VERSION : 0.0
   STRUCT
      Config_bit_Converter : Bool;   // Configuration with frequency converter
      Config_bit_Converter_SW : Bool;   // Configuration with frequency converter with Set value
      Config_bit_Heating_ON : Bool;
      config_bit_Heating_Int : Bool;
      Config_bit_Cooling_ON : Bool;
      Config_bit_Cooling_Int : Bool;
      Config_bit_Filling_ON : Bool;
      Config_bit_Filling_Int : Bool;
      Config_bit_Charging_ON : Bool;
      Config_bit_Charging_Int : Bool;
      RunTime : S5Time;
      PauseTime : S5Time;
   END_STRUCT;
END_TYPE

TYPE "UDT102_RefillingState"
TITLE = State of refilling tank
VERSION : 0.0
   STRUCT
      Value_No : Int;   // Storage of shot amout if refilling after shot amount reached is selected
      Fault_Exist : Bool;   // A fault inside this function exist
      FaultLevel_1 : Bool;   // A fault level 1 inside this function exist
      FaultLevel_2 : Bool;   // A fault level 2 inside this function exist
      FaultLevel_3 : Bool;   // A fault level 3 inside this function exist
      Spare_1_5 : Bool;
      Spare_1_6 : Bool;
      Select_refilling : Bool;   // Requirement of refilling the tank
      Spare_2_0 : Bool;
      Spare_2_1 : Bool;
      Spare_2_2 : Bool;
      Ramp_MH_open : Bool;   // Flag to compare if refilling after shot amount reached is selected
      FLT_Alarm_N2 : Bool;   // Fault alarm nitrogen at tank (1)
      Preagitation_runs : Bool;   // Pre mixing time before refilling the tank
      Filling_Start : Bool;   // Pre mixing time finished -> start refilling the tank
      Fillingtime_runs : Bool;   // Tank refilling started and refillingtime monitoring active
      Select_Filling_with_Time : Bool;   // Requirement of refilling the tank after time ("IN_Zeit_bis_Bef" >0)
      Block_is_activ : Bool;   // The funktion block passed through // Info min. 1 tank active
      Max_Level : Bool;   // Level of Tank over maximum
      Stop_Level_Filling : Bool;   // Level of Tank over filling level
      Start_Level_Filling : Bool;   // Level of Tank beneath filling level
      Min_Level : Bool;   // Level of Tank beneath mimimum
      Enable_Agitator : Bool;   // Level of Tank for enabling agitator
      Switch_Refilling_ON_OFF : Bool;   // Switch refilling ON/OFF (external Signal)
      ButtonLeakageMonitorOFF : Bool;   // Button bridging leakage monitoring
      PreWarning_Min_Level : Bool;   // Level of Tank reached pre warnings
      Switch_DrainTank_ON_OFF : Bool;   // Switch drain tank ON/OFF (external Signal)
      LevelTriptray : Bool;   // Level Triptry was detected
      Switch_Refilling_from_Barrel_ON_OFF : Bool;   // Anwahl des Befüllventils durch Faßstation
      Spare_5_4 : Bool;
      Spare_5_5 : Bool;
      Spare_5_6 : Bool;
      Spare_5_7 : Bool;
      State_Refilling : Int;   // 1->Refilling ON; 2->Fault Refilling; 3->Refilling requested but not on
   END_STRUCT;
END_TYPE

TYPE "UDT100_AggitatorState"
TITLE = State of auxiliary drive
VERSION : 0.0
   STRUCT
      FLT_Exist : Bool;
      MES_Run_Heating : Bool;
      MES_Run_Cooling : Bool;
      MES_Run_Filling : Bool;
      MES_Run_Charging : Bool;
      FaultLevel_3 : Bool;   // A fault group 3 exist
      Spare0_7 : Bool;
      Reset_Intervall : Bool;   // Reset of intervall- mode at running- and pausetime
      Run : Bool;   // Drive at intervall- mode in running
      Pause : Bool;   // Drive at intervall- mode in pause time
      No_Pausetime : Bool;   // Running- or pausetime is "0" -> drive is running continuously
      Ramp_CVoltage_Off : Bool;   // Flag of delay to switch ON after power lost
      Start_Startupdelay : Bool;   // Information delay time to switch ON after power lost is running
      Disable_Start : Bool;   // Information delay time to switch ON after power lost is running
      Switch_Drive_ON_OFF : Bool;   // Switch auxiliary drive ON-OFF (external signal)
      State_Drive : Int;   // 1->Drive ON; 2->Fault Drive; 3->Drive requested but not on
   END_STRUCT;
END_TYPE

TYPE "UDT101_auxiDriveState"
TITLE = State of auxiliary drive
VERSION : 0.0
   STRUCT
      FLT_Motorprotection : Bool;   // Fault: Powersupply or motorprotection of drive
      FLT_FC : Bool;   // Fault: Frequncyconverter of drive is faulty
      FLT_MaxP_MaxLTripTray : Bool;   // Fault: Maximium component pressure or maximum filling level triptray exceeded
      FLT_Dryrunsafety : Bool;   // Fault: Dry running of drive activated
      FLT_wrong_Timevalue : Bool;   // Information a time value was inputed, which makes no sense
      FLT_MaxPressureDiff : Bool;   // Fault: Max. pressure difference at filter
      FLT_MotorFan : Bool;   // Fault: Motorprotection external fan of motor
      FaultExist : Bool;   // A fault message exist
      Reset_Intervall : Bool;   // Reset of intervall- mode at running- and pausetime
      Run : Bool;   // Drive at intervall- mode in running
      Pause : Bool;   // Drive at intervall- mode in pause time
      No_Pausetime : Bool;   // Running- or pausetime is "0" -> drive is running continuously
      Ramp_CVoltage_Off : Bool;   // Flag of delay to switch ON after power lost
      Start_Startupdelay : Bool;   // Information delay time to switch ON after power lost is running
      Disable_Start : Bool;   // Information delay time to switch ON after power lost is running
      Switch_Drive_ON_OFF : Bool;   // Switch auxiliary drive ON-OFF (external signal)
      State_Drive : Int;   // 1->Drive ON; 2->Fault Drive; 3->Drive requested but not on
      Config_bit_normal : Bool;   // Drive config as agitator, heatexchanger or circulationpump -> normal (agitator)
      Config_bit_char : Bool;   // Drive config as circulation pump and filling pump
      config_bit_feed : Bool;   // Drive config as circulation pump and feed pump
      Config_bit_split : Bool;   // Drive config as edge filter
      Config_bit_with_FC : Bool;   // Drive config as with frequency unit for example as agitator
      Config_bit_5 : Bool;
      Config_bit_6 : Bool;
      Config_bit_7 : Bool;
      Spare_5_0 : Bool;
      Spare_5_1 : Bool;
      Spare_5_2 : Bool;
      Spare_5_3 : Bool;
      Spare_5_4 : Bool;
      Spare_5_5 : Bool;
      Spare_5_6 : Bool;
      Spare_5_7 : Bool;
   END_STRUCT;
END_TYPE

TYPE "UDT105_Controller_State"
TITLE = State of 2-point controller tempering
VERSION : 0.1
   STRUCT
      CoolingActive : Bool;
      HeatingActive : Bool;
      CoolingRequest : Bool;
      HeatingRequest : Bool;
      FLT_Fuse_Heating : Bool;
      HF_Set_Cooling : Bool;
      HF_Set_Heating : Bool;
      Spare_13 : Bool;
      Trigger : Bool;   // Trigger to start calculation pulstime
      Start_delay_puls : Bool;
      Fault_Exist : Bool;
      Spare_1_3 : Bool;
      Spare_1_4 : Bool;
      Spare_1_5 : Bool;
      Spare_1_6 : Bool;
      Switch_Temp_ON_OFF : Bool;
      PulsTime : DInt;   // Time to switch on valve heatexchanger
      State_Temp : Int;
   END_STRUCT;
END_TYPE

TYPE "UDT106_Vacuum_Status"
TITLE = State of vacuum unit
VERSION : 0.1
   STRUCT
      Spare_0_0 : Bool;
      Spare_0_1 : Bool;
      Switch_Vacuum_ON_OFF : Bool;   // Switch auxiliary drive ON-OFF (external signal)
      Spare_0_2 : Bool;
      Spare_0_4 : Bool;
      Spare_0_5 : Bool;
      Spare_0_6 : Bool;
      Spare_0_7 : Bool;
      FLT_PVacuum : Bool;   // Pressure vacuum not reached
      Spare_1_1 : Bool;
      Spare_1_2 : Bool;
      Spare_1_3 : Bool;
      Spare_1_4 : Bool;
      Spare_1_5 : Bool;
      Spare_1_6 : Bool;
      Spare_1_7 : Bool;
      Status_Vacuum : Int;   // 1->Drive ON; 2->Fault Drive; 3->Drive requested but not on
   END_STRUCT;
END_TYPE

TYPE "UDT107_MicroMeteringUnit"
TITLE = State of micro metering unit
VERSION : 0.0
   STRUCT
      FLT_MultibleAllocation : Bool;   // Allocation of metering unit at more then one connector
      FLT_NotSelected : Bool;   // Selection of metering unit by switch missing
      FLT_PowerSupply : Bool;   // Power supply metering unit faulty
      FLT_Watchdog : Bool;   // No sign of live signal from metering unit
      FLT_NotOperative : Bool;   // Metering unit not ready for operation
      FLT_NotAllocated : Bool;   // Metering unit not allocated to mixinghead connector
      Spare01 : Bool;
      Spare02 : Bool;
      ReleaseMH : Bool;   // Release mixing head
      Spare_1_1 : Bool;   // Flag of delay to switch ON after power lost
      Enableclosedloop : Bool;   // PLC-release to control the component flow at modul
      Metering_to_PUC : Bool;   // Request of metering the component
      Flag_QPB : Bool;   // Flag of the signal to switch over to the quick pressure build up
      StartQPB : Bool;   // Signal start quick pressure build up
      Switch_Drive_ON_OFF : Bool;   // Switch micro metering unit ON-OFF (external signal)
      Spare_1_7 : Bool;
      State_Drive : Int;   // 1->Drive ON; 2->Fault Drive; 3->Drive requested but not on
      ConnectionPlace : Array[1..16] of Bool;   // Possible places to connect a metering unit
      AllocConnectPlaceNo : Int;   // Allocation metering unit at mixighead connector (place no at mixingheads)
   END_STRUCT;
END_TYPE

TYPE "UDT108_AbortComponent"
VERSION : 0.1
   STRUCT
      Spare_0_0 : Bool;
      Spare_0_1 : Bool;
      Abort_ON_OFF : Bool;   // Switch auxiliary device ON-OFF (external signal)
      Spare_0_2 : Bool;
      Spare_0_4 : Bool;
      Spare_0_5 : Bool;
      Spare_0_6 : Bool;
      Spare_0_7 : Bool;
      Spare_1_0 : Bool;
      Spare_1_1 : Bool;
      Spare_1_2 : Bool;
      Spare_1_3 : Bool;
      Spare_1_4 : Bool;
      Spare_1_5 : Bool;
      Spare_1_6 : Bool;
      Spare_1_7 : Bool;
      Status_Abort : Int;   // 1->Drive ON; 2->Fault Drive; 3->Drive requested but not on
   END_STRUCT;
END_TYPE

TYPE "UDT103_RefilStationState"
TITLE = State of material container (storage unit)
VERSION : 0.1
   STRUCT
      Message_No_Drum : Bool;   // Meldung: Es ist kein Faß in der Containerstation vorhanden
      Message_DrumExist : Bool;
      FLT_Min_Pressure_Air : Bool;   // Störung: Eingestellter min. Druck der Luftversorgung unterschritten
      FLT_MinPressureAirPump : Bool;   // Störung: Das Faß in der Containerstation ist leer! Bitte wechseln!
      FLT_Heat : Bool;   // Störung: Der Trockenlaufschutz an der Kreislaufpumpe hat angesprochen
      FLT_Spare05 : Bool;   // Störung: Der Komponentendruck in der Kreislaufleitung wurde überschritten
      FLT_Spare06 : Bool;
      FLT_Spare07 : Bool;
      Agitator_before_Fill_DT : Bool;   // Rührwerk: Toggelbit zum Ansteuern des Rührwerkes vor der Befüllung des TB
      Agitator_after_Fill_Cont : Bool;   // Rührwerk: Toggelbit zum Ansteuern des Rührwerkes nach der Befüllung des Cont
      Filling_Cont_start : Bool;   // Befüllung: Befüllung des Containers starten
      Filling_Cont_Puls_stop : Bool;   // Befüllung: Impulsmerker für das stoppen der Befüllung
      Filling_Cont_Started : Bool;   // Befüllung: Die Befüllung des Containers wurde gestartet
      Filling_Cont_Drum_empty : Bool;   // Befüllung: Das Signal für "MLD Faß leer" kann ausgewertet werden
      Filling_Cont_MaxFilltime : Bool;   // Befüllung: Die Füllzeit des Containers wurde überschritten
      Filling_Cont_Spare_2_5 : Bool;
      Agitator_Cont_PreAgit : Bool;   // Rührwerk: Aufrühren des Rührwerkes des Contaioners
      Agitator_Cont_Puls_Start : Bool;   // Rührwerk: Impulsmerker für das Starten des Rührwerkes
      Agitator_Cont_Runtim_End : Bool;   // Rührwerk: Laufzeit des Rührwerkes ist abgelaufen
      Agitator_Cont_Release_DT : Bool;   // Rührwerk: Vorrührzeit ist beendet -> Freigabe zum Befüllen des Tagesbehälters
      Agitator_Cont_Release : Bool;
      RCL_Cont_Puls_Start : Bool;   // Kreislaufpumpe: Impulsmerker für das Starten der Kreislaufpumpe
      RCL_Cont_Dryprotection : Bool;   // Kreislaufpumpe: Einschaltverzögerung des Trockenlaufschutzes ist aktiviert
      RCL_Cont_Runtime_Ende : Bool;   // Kreislaufpumpe: Laufzeit der Kreislaufpumpe ist abgelaufen
      RCL_Cont_Release_Fill_DT : Bool;   // Kreislaufpumpe: Freigabesignal für die Befüllung des Tagesbehälters
      RCL_Cont_Spare_3_7 : Bool;
      Agitator : "UDT101_auxiDriveState";
      Pump : "UDT101_auxiDriveState";
      Filling : "UDT102_RefillingState";
      Switch_ONOFF_Heat01 : Bool;
      Switch_ONOFF_Heat02 : Bool;
      State_Heat1 : Int;   // 1-> ON; 2->Fault; 3->Requested but not on
      State_Heat2 : Int;   // 1-> ON; 2->Fault; 3->Requested but not on
   END_STRUCT;
END_TYPE

TYPE "UDT2002_Output_Faurecia"
VERSION : 0.1
   STRUCT
      Machinestatus : Struct
         AUTO : Bool := FALSE;   // 1 = machine is in Automatic and ready for production
         MANUAL : Bool := FALSE;   // 1 = machine is in Manual mode
         SERVICE : Bool := FALSE;   // 0 = machine is in Service mode (only simulated shots, no mixhead opening)
         CYCLE_RUN : Bool := FALSE;   // 1 = foam cycle is active
         READY : Bool := FALSE;   // 1 = waiting for shot release
         POURING : Bool := FALSE;   // 1 = shot is running (also a "service shot")
         SHOTEND : Bool := FALSE;   // 1 = Shot is done
         CPFORWARD : Bool := FALSE;   // 1 = Cleaning piston is in cleaning position
         FAULTGROUP1 : Bool := FALSE;   // 0 = machine is faulted (only group 1)
         Startbutton : Bool := FALSE;   // 1 = Pad control STARTSHOT push button
         Kreislauf : Bool := FALSE;   // 1 = machine is in reduced circulation
         ACK : Bool := FALSE;   // Acknowledge foam parameters
         Reserve5 : Bool := FALSE;
         Reserve6 : Bool := FALSE;
         Reserve7 : Bool := FALSE;
         Watchdog : Bool := FALSE;
      END_STRUCT;
      Act_Comp_Values : Struct
         Flow_C1 : Word := W#16#0;   // Actual flow C1 in 1/10g/s
         Flow_C2 : Word := W#16#0;   // Actual flow C2 in 1/10g/s
         mixingratio : Word := W#16#0;   // ISO Mixingratio, POLY=100%
         Feedline_Pressure_C1 : Word := W#16#0;   // Actual pressure feedline C1 in 1/10 bar
         Feedline_Pressure_C2 : Word := W#16#0;   // Actual pressure feedline C2 in 1/10 bar
         MH_Pressure_C1 : Word := W#16#0;   // Mixhead pressure (Option) in 1/10 bar
         MH_Pressure_C2 : Word := W#16#0;   // Mixhead pressure (Option) in 1/10 bar
         Tank_Temp_C1 : Word := W#16#0;   // in 1/10°C
         Tank_Temp_C2 : Word := W#16#0;   // in 1/10°C
         MH_Temp_C1 : Word := W#16#0;   // Mixhead Temp (Option) in 1/10°C
         MH_Temp_C2 : Word := W#16#0;   // Mixhead Temp (Option) in 1/10°C
      END_STRUCT;
      Last_Shot_datas : Struct
         shottime : DWord := DW#16#0;   // in ms
         Flow_C1 : Word := W#16#0;   // in 1/10g/s
         Flow_C2 : Word := W#16#0;   // in 1/10g/s
         mixingratio : Word := W#16#0;   // ISO Mixingratio, POLY=100%
         weight : Word := W#16#0;   // last shot weight in 1/10 g
         Feedline_Pressure_C1 : Word := W#16#0;   // in 1/10bar
         Feedline_Pressure_C2 : Word := W#16#0;   // in 1/10bar
         MH_Pressure_C1 : Word := W#16#0;   // Mixhead pressure (Option) in 1/10bar
         MH_Pressure_C2 : Word := W#16#0;   // Mixhead pressure (Option) in 1/10bar
         MH_Temp_C1 : Word := W#16#0;   // Mixhead Temp (Option) in 1/10°C
         MH_Temp_C2 : Word := W#16#0;   // Mixhead Temp (Option) in 1/10°C
      END_STRUCT;
      Reserve : Struct
         Reserve1 : Word;
         Reserve2 : Word;
      END_STRUCT;
      Alarm_GRP1_1 : Array[0..15] of Bool;   // n+48
      Alarm_GRP1_2 : Array[0..15] of Bool;   // n+50
      Alarm_GRP1_3 : Array[0..15] of Bool;   // n+52
      Alarm_GRP1_4 : Array[0..15] of Bool;   // n+54
      Alarm_GRP1_5 : Array[0..15] of Bool;   // n+56
      Alarm_GRP1_6 : Array[0..15] of Bool;   // n+58
      Alarm_GRP1_7 : Array[0..15] of Bool;   // n+60
      Alarm_GRP1_8 : Array[0..15] of Bool;   // n+62
      Alarm_GRP1_9 : Array[0..15] of Bool;   // n+64
      Alarm_GRP1_10 : Array[0..15] of Bool;   // n+66
      Alarm_GRP1_11 : Array[0..15] of Bool;   // n+68
      Alarm_GRP1_12 : Array[0..15] of Bool;   // n+70
      Alarm_GRP1_13 : Array[0..15] of Bool;   // n+72
      Alarm_GRP1_14 : Array[0..15] of Bool;   // n+74
      Alarm_GRP1_15 : Array[0..15] of Bool;   // n+76
      Alarm_GRP1_16 : Array[0..15] of Bool;   // n+78
      Alarm_GRP2_1 : Array[0..15] of Bool;   // n+80
      Alarm_GRP2_2 : Array[0..15] of Bool;   // n+82
      Alarm_GRP2_3 : Array[0..15] of Bool;   // n+84
      Alarm_GRP2_4 : Array[0..15] of Bool;   // n+86
      Alarm_GRP3_1 : Array[0..15] of Bool;   // n+88
      Alarm_GRP3_2 : Array[0..15] of Bool;   // n+90
      Alarm_GRP3_3 : Array[0..15] of Bool;   // n+92
      Alarm_GRP3_4 : Array[0..15] of Bool;   // n+94
      Alarm_GRP3_5 : Array[0..15] of Bool;   // n+96
      Alarm_GRP3_6 : Array[0..15] of Bool;   // n+98
      Alarm_GRP3_7 : Array[0..15] of Bool;   // n+100
      Alarm_GRP3_8 : Array[0..15] of Bool;   // n+102
      Alarm_GRP3_9 : Array[0..15] of Bool;   // n+104
      Alarm_GRP3_10 : Array[0..15] of Bool;   // n+106
      Alarm_GRP3_11 : Array[0..15] of Bool;   // n+108
      Alarm_GRP3_12 : Array[0..15] of Bool;   // n+110
      Alarm_GRP3_13 : Array[0..15] of Bool;   // n+112
      Alarm_GRP3_14 : Array[0..15] of Bool;   // n+114
      Alarm_GRP3_15 : Array[0..15] of Bool;   // n+116
      Alarm_GRP3_16 : Array[0..15] of Bool;   // n+118
      Alarm_GRP3_17 : Array[0..15] of Bool;   // n+120
      Alarm_GRP3_18 : Array[0..15] of Bool;   // n+122
      Alarm_GRP3_19 : Array[0..15] of Bool;   // n+124
      Alarm_GRP3_20 : Array[0..15] of Bool;   // n+126
      Alarm_GRP3_21 : Array[0..15] of Bool;   // n+128
      Alarm_GRP3_22 : Array[0..15] of Bool;   // n+130
      Alarm_GRP3_23 : Array[0..15] of Bool;   // n+132
      Alarm_GRP3_24 : Array[0..15] of Bool;   // n+134
      Alarm_GRP3_25 : Array[0..15] of Bool;   // n+136
      Alarm_GRP3_26 : Array[0..15] of Bool;   // n+138
      Alarm_GRP3_27 : Array[0..15] of Bool;   // n+140
      Alarm_GRP3_28 : Array[0..15] of Bool;   // n+142
      Message_1 : Array[0..15] of Bool;   // n+144
      Message_2 : Array[0..15] of Bool;   // n+146
      Message_3 : Array[0..15] of Bool;   // n+148
      Message_4 : Array[0..15] of Bool;   // n+150
      Message_5 : Array[0..15] of Bool;   // n+152
      Message_6 : Array[0..15] of Bool;   // n+154
      Message_7 : Array[0..15] of Bool;   // n+156
      Message_8 : Array[0..15] of Bool;   // n+158
      Message_9 : Array[0..15] of Bool;   // n+160
      Message_10 : Array[0..15] of Bool;   // n+162
   END_STRUCT;
   // // Alarm_GRP1_1[8] : " Operating mode changed during foam cycle "
   // // Alarm_GRP1_1[9] : " Shottime too small"
   // // Alarm_GRP1_1[10] : " No COU selected "
   // // Alarm_GRP1_1[11] : " Selected COU not valid "
   // // Alarm_GRP1_1[12] : " Maximum-shot-time overstepped "
   // // Alarm_GRP1_1[0] : Machine start a new program without ends the existing
   // // Alarm_GRP1_1[1] : Machine reset the program number during shot
   // // Alarm_GRP1_1[2] : " Wrong Mixinghead-Number assigned in the foam program "
   // // Alarm_GRP1_1[3] : No foaming program selected
   // // Alarm_GRP1_1[4] : " Mixinghead doesn't open"
   // // Alarm_GRP1_1[5] : " Mixinghead doesn't close "
   // // Alarm_GRP1_1[6] : Mixinghead open without control
   // // Alarm_GRP1_1[7] : Mixinghead close during shot
   // // Alarm_GRP1_2[8] : Shot aborted
   // // Alarm_GRP1_2[9] : Mixinghead bouncing during control
   // // Alarm_GRP1_2[10] : General fault from PUC
   // // Alarm_GRP1_2[13] : " Fault alien plant interface 1"
   // // Alarm_GRP1_2[15] : " Profibus module machine faulty (DP:3) "
   // // Alarm_GRP1_2[0] : " ET200 profibus module faulty"
   // // Alarm_GRP1_2[6] : " Maximum-pressure component Poly
   // // Alarm_GRP1_2[7] : " Maximum-pressure component Iso
   // // Alarm_GRP1_3[10] : " Tolerance + pressure Poly at Mixinghead 1"
   // // Alarm_GRP1_3[11] : " Tolerance + pressure Iso at Mixinghead 1"
   // // Alarm_GRP1_3[0] : " Min.-pressure component Poly
   // // Alarm_GRP1_3[1] : " Min.-pressure component Iso
   // // Alarm_GRP1_3[4] : " Tolerance - pressure Poly at Mixinghead 1"
   // // Alarm_GRP1_3[5] : " Tolerance - pressure Iso at Mixinghead 1"
   // // Alarm_GRP1_4[10] : " Tank pressure is missing Poly
   // // Alarm_GRP1_4[11] : " Tank pressure is missing Iso
   // // Alarm_GRP1_4[4] : " Min.-level tank Poly
   // // Alarm_GRP1_4[5] : " Min.-level tank Iso
   // // Alarm_GRP1_5[8] : " Tolerance - tank temperature Poly
   // // Alarm_GRP1_5[9] : " Tolerance - tank temperature Iso
   // // Alarm_GRP1_5[14] : " Max.Level tank Poly
   // // Alarm_GRP1_5[15] : " Max.Level tank Iso
   // // Alarm_GRP1_5[2] : " Tolerance + tank temperature Poly
   // // Alarm_GRP1_5[3] : " Tolerance + tank temperature Iso
   // // Alarm_GRP1_6[8] : " Drip-tray full Poly
   // // Alarm_GRP1_6[9] : " Drip-tray full Iso
   // // Alarm_GRP1_6[12] : " Tolerance - flow Poly
   // // Alarm_GRP1_6[13] : " Tolerance - flow Iso
   // // Alarm_GRP1_6[0] : " Tolerance + flow Poly
   // // Alarm_GRP1_6[1] : " Tolerance + flow Iso
   // // Alarm_GRP1_6[4] : " Tolerance - MR Poly
   // // Alarm_GRP1_6[5] : " Tolerance - MR Iso
   // // Alarm_GRP1_7[8] : " Tolerance + MR Poly
   // // Alarm_GRP1_7[9] : " Tolerance + MR Iso
   // // Alarm_GRP1_7[12] : " Motor-protection Mixinghead-Hydraulic "
   // // Alarm_GRP1_7[13] : " Maximum-temperature oil Mixinghead-Hydraulic "
   // // Alarm_GRP1_7[14] : " Min.level oil Mixinghead-Hydraulic"
   // // Alarm_GRP1_7[15] : " Maximum-contact not reached Mixinghead-Hydraulic "
   // // Alarm_GRP1_7[6] : " Motor-protection pump Poly
   // // Alarm_GRP1_7[7] : " Motor-protection pump Iso
   // // Alarm_GRP1_8[10] : " Tolerance - temperature Poly at Mixinghead 1"
   // // Alarm_GRP1_8[11] : " Tolerance - temperature Iso at Mixinghead 1"
   // // Alarm_GRP1_8[0] : " Fault fequency converter pump Poly
   // // Alarm_GRP1_8[1] : " Fault fequency converter pump Iso
   // // Alarm_GRP1_8[4] : " Tolerance + temperature Poly at Mixinghead 1"
   // // Alarm_GRP1_8[5] : " Tolerance + temperature Iso at Mixinghead 1"
   // // Alarm_GRP1_10[14] : " Motor-protection feeding pump Poly
   // // Alarm_GRP1_10[15] : " Motor-protection feeding pump Iso
   // // Alarm_GRP1_11[2] : " Maximum runtime reached feeding pump Poly "
   // // Alarm_GRP1_11[3] : " Maximum runtime reached feeding pump Iso "
   // // Alarm_GRP2_1[8] : " Fault Alien plant"
   // // Alarm_GRP2_1[12] : " Min.level tank Poly during Cycle"
   // // Alarm_GRP2_1[13] : " Min.level tank Iso during Cycle"
   // // Alarm_GRP2_1[7] : " Drip-tray full Iso during cycle"
   // // Alarm_GRP2_1[6] : " Drip-tray full Poly during cycle"
   // // Alarm_GRP2_3[10] : " Pre-warning maximum-temperature mixingheadhydraulic"
   // // Alarm_GRP3_1[8] : " Motor-protection circulating pump/agitator Poly"
   // // Alarm_GRP3_1[9] : " Motor-protection circulating pump/agitator Iso
   // // Alarm_GRP3_1[2] : " Fault FC agitator Poly"
   // // Alarm_GRP3_1[3] : " Fault FC agitator Iso
   // // Alarm_GRP3_2[12] : " Filling time exceeded tank Poly"
   // // Alarm_GRP3_2[13] : " Filling time exceeded tank Iso
   // // Alarm_GRP3_2[0] : " Level sensor faulty Poly"
   // // Alarm_GRP3_2[1] : " Level sensor faulty Iso
   // // Alarm_GRP3_2[7] : " Max.Level tank Iso
   // // Alarm_GRP3_2[6] : " Max.Level tank Poly
   // // Alarm_GRP3_3[11] : " Pre-mixing station is not ready"
   // // Alarm_GRP3_3[0] : " Motor-protection split-filter Poly
   // // Alarm_GRP3_3[1] : " Motor-protection split-filter Iso
   // // Alarm_GRP3_4[10] : " Oil filter contaminated Mixinghead hydraulic"
   // // Alarm_GRP3_4[11] : " Oil filter contaminated Mixinghead hydraulic (High pressure) "
   // // Alarm_GRP3_5[15] : " Maximum-waiting time after circulation time 1 "
   // // Alarm_GRP3_5[14] : " No cycle time programmed "
   // // Alarm_GRP3_5[0] : n+96
   // // Alarm_GRP3_5[2] : " Fault Fuse"
   // // Alarm_GRP3_5[3] : " Fault air-dryer "
   // // Alarm_GRP3_5[4] : " Fault heat-balancing unit "
   // // Alarm_GRP3_5[5] : " Fault heating supply "
   // // Alarm_GRP3_5[7] : " Fault Alien plant"
   // // Alarm_GRP3_6[8] : " Fault hose-heating Poly"
   // // Alarm_GRP3_6[9] : " Fault hose-heating Iso"
   // // Alarm_GRP3_6[10] : " Fault mixinghead heating"
   // // Alarm_GRP3_6[14] : " Fault Parity bit Alien plant 1"
   // // Alarm_GRP3_6[15] : " Fault Parity bit Alien plant 2"
   // // Alarm_GRP3_6[2] : " Closed loop metering limit reached Poly
   // // Alarm_GRP3_6[3] : " Closed loop metering limit reached Iso
   // // Alarm_GRP3_11[8] : " Profibus module Mixinghead 1 faulty "
   // // Alarm_GRP3_11[9] : " Profibus module Mixinghead 2 faulty "
   // // Alarm_GRP3_12[15] : " Profibus connection to robot faulty"
   // // Alarm_GRP3_12[0] : " Profibus connection to container-station faulty"
   // // Alarm_GRP3_12[1] : " Profibus-connection to alien plant faulty"
   // // Alarm_GRP3_13[0] : " Cleaning-plunger too slow MH1 "
   // // Alarm_GRP3_13[1] : " Cleaning-plunger leaves rear position during shot MH1"
   // // Alarm_GRP3_13[2] : " No cleaning-plunger initiator MH1"
   // // Alarm_GRP3_13[3] : " Cleaning-plunger too slow MH2 "
   // // Alarm_GRP3_13[4] : " Cleaning-plunger leaves rear position during shot MH2"
   // // Alarm_GRP3_13[5] : " No cleaning-plunger initiator MH2"
   // // Alarm_GRP3_16[2] : " Fault nucleation unit Poly "
   // // Alarm_GRP3_16[3] : " Fault nucleation unit Iso "
   // // Alarm_GRP3_17[10] : " Timeout during fast pressure build up (FPB)"
   // // Alarm_GRP3_17[12] : " Min material-level flushing-agent pump"
   // // Alarm_GRP3_17[5] : " Warning - pressure Poly at MH 1"
   // // Alarm_GRP3_17[6] : " Warning - pressure Iso at MH 1"
   // // Alarm_GRP3_18[9] : " Warning + pressure Poly at MH 1"
   // // Alarm_GRP3_18[10] : " Warning + pressure Iso at MH 1"
   // // Alarm_GRP3_18[13] : " Warning - temperature Poly at MH 1"
   // // Alarm_GRP3_18[14] : " Warning - temperature Iso at MH 1"
   // // Alarm_GRP3_18[1] : " Warning + temperature Poly at MH 1"
   // // Alarm_GRP3_18[2] : " Warning + temperature Iso at MH 1"
   // // Alarm_GRP3_18[5] : " Warning - flow Poly
   // // Alarm_GRP3_18[6] : " Warning - flow Iso
   // // Alarm_GRP3_19[9] : " Warning + flow Poly
   // // Alarm_GRP3_19[10] : " Warning + flow Iso
   // // Alarm_GRP3_19[13] : " Warning - MR Poly
   // // Alarm_GRP3_19[14] : " Warning - MR Iso
   // // Alarm_GRP3_19[1] : " Warning + MR Poly
   // // Alarm_GRP3_19[2] : " Warning + MR Iso
   // // Alarm_GRP3_19[5] : " Warning - shottime Mixinghead 1"
   // // Alarm_GRP3_19[6] : " Warning + shottime Mixinghead 1"
   // // Alarm_GRP3_19[7] : " Warning - weight Mixinghead 1"
   // // Alarm_GRP3_20[8] : " Warning + weight Mixinghead 1"
   // // Alarm_GRP3_20[9] : " Warning - temperature tank Poly
   // // Alarm_GRP3_20[10] : " Warning - temperature tank Iso
   // // Alarm_GRP3_20[13] : " Warning + temperature tank Poly
   // // Alarm_GRP3_20[14] : " Warning + temperature tank Iso
   // // Alarm_GRP3_21[2] : " System-fault robot"
   // // Alarm_GRP3_23[11] : " Supply-fault robot cabinet"
   // // Alarm_GRP3_24[3] : " Interval time too short"
   // // Message_1[8] : " No control voltage "
   // // Message_1[9] : " Container-station fault"
   // // Message_1[10] : " ESTOP machine "
   // // Message_1[11] : " EMERGENCY STOP machine 2"
   // // Message_1[12] : " EMERGENCY HALT (Safety gate?)"
   // // Message_1[13] : " ESTOP nucleation unit "
   // // Message_1[15] : " ESTOP user panel "
   // // Message_1[0] : " ESTOP Pentanstation"
   // // Message_1[1] : " ESTOP mould carrier"
   // // Message_1[2] : " ESTOP robot"
   // // Message_1[3] : " ESTOP alien plant interface"
   // // Message_2[6] : " EMERGENCY STOP on container-station"
   // // Message_3[8] : " ESTOP user panel mixinghead 1"
   // // Message_3[9] : " ESTOP user panel mixinghead 2"
   // // Message_6[15] : " Weekend mode is active"
   // // Message_6[4] : " Robot not in Auto mode"
   // // Message_9[11] : " Start-up delay of FCs is running, please wait"
END_TYPE

TYPE "UDT111_GenAuxDrivesState"
TITLE = State of additional drives (please customize)
VERSION : 0.1
   STRUCT
      FanHousing : "UDT101_auxiDriveState";
      AuxDriveState_Spare01 : "UDT101_auxiDriveState";
      AuxDriveState_Spare02 : "UDT101_auxiDriveState";
      AuxDriveState_Spare03 : "UDT101_auxiDriveState";
      AuxDriveState_Spare04 : "UDT101_auxiDriveState";
      AuxDriveState_Spare05 : "UDT101_auxiDriveState";
      AuxDriveState_Spare06 : "UDT101_auxiDriveState";
      AuxDriveState_Spare07 : "UDT101_auxiDriveState";
      AuxDriveState_Spare08 : "UDT101_auxiDriveState";
      AuxDriveState_Spare09 : "UDT101_auxiDriveState";
      AuxDriveState_Spare10 : "UDT101_auxiDriveState";
   END_STRUCT;
END_TYPE

TYPE "UDT109_CoverLift"
TITLE = State of cover lift
VERSION : 0.1
   STRUCT
      Spare_0_0 : Bool;
      Spare_0_1 : Bool;
      Switch_ON_OFF : Bool;   // Switch auxiliary drive ON-OFF (external signal)
      Spare_0_2 : Bool;
      CoverReadyToClose : Bool;   // Cover ready to close at tank
      Spare_0_5 : Bool;
      Spare_0_6 : Bool;
      Spare_0_7 : Bool;
      FLT_P_Air : Bool;   // Pressure vacuum not reached
      FLT_LiftingTooSlow : Bool;   // Monitoring time lifting exceeded
      FLT_DropingTooSlow : Bool;   // Monitoring time droping exceeded
      Spare_1_3 : Bool;
      Spare_1_4 : Bool;
      Spare_1_5 : Bool;
      Spare_1_6 : Bool;
      Spare_1_7 : Bool;
      Status : Int;   // 1->Drive ON; 2->Fault Drive; 3->Drive requested but not on
   END_STRUCT;
END_TYPE

TYPE "ABB_IRC5_Status"
TITLE = Signals interface robot
VERSION : 0.0
   STRUCT
      Auto_mode_requested : Bool;   // Automatic mode requested
      Manual_mode_requested : Bool;   // Manual mode requested
      Auto_accepted : Bool;   // Automatic accepted
      Freigabe_Schaeumzyklus : Bool;   // Release foaming
      Release_foaming : Bool;   // Start foaming cycle
      Shot_time_received : Bool;   // Shot time received
      Data_transmitted : Bool;   // Data transmitted
      Data_inv_transmitted : Bool;   // Data inverse transmitted
      Interface_OK : Bool;   // Interface OK
      STG_System : Bool;   // Fault from system
      Fault_from_system : Bool;   // Fault from interface
      Fault_observed : Bool;   // Fault observed
      Escape_program : Bool;   // Escape program
      Motion_prog01_existing : Bool;   // Motion program 1 existing
      Motion_prog02_existing : Bool;   // Motion program 2 existing
      Motion_prog03_existing : Bool;   // Motion program 3 existing
      Robot_ProgNo_Mould_1 : Byte;   // Roboter program number mould 1
      Robot_ProgNo_Mould_2 : Byte;   // Roboter program number mould 2
      Robot_ProgNo_Mould_3 : Byte;   // Roboter program number mould 3
      Robot_processing_prog : Bool;   // Roboter processing program
      HFShotDigOut_open_MH : Bool;
      doShotDigOut_open_MH : Bool;
      HF_next_partshot : Bool;   // Flankenhilfsmerker für die Ermittlung eines neuen Verfahrprogramms // Teilschuß
      HF_Robot_not_in_Auto : Bool;   // Flankenhilfsmerker für das zurücksetzten des Signals "Roboter nicht in Auto"
      Robot_not_in_Auto : Bool;   // Roboter not in automatic mode
      Start_Synchronization : Bool;
      FLT_SyncPosition : Bool;   // Robot will perform the synchronization
      FHM_SyncEPS : Bool;   // The Synchronization position is not correct
      CleaningSelected : Bool;   // Flag for the information that a cleaning was selected
      CleaningActiv : Bool;   // Flag for the information that a cleaning is activ
      FHM_CleaningActiv : Bool;   // Helpflag for the information that a cleaning is activ
      Reserve_6_4 : Bool;
      Reserve_6_5 : Bool;
      Reserve_6_6 : Bool;
      Reserve_6_7 : Bool;
      Reserve_7_0 : Bool;
      Reserve_7_1 : Bool;
      Reserve_7_2 : Bool;
      Reserve_7_3 : Bool;
      Reserve_7_4 : Bool;
      Reserve_7_5 : Bool;
      Reserve_7_6 : Bool;
      Reserve_7_7 : Bool;
      Reserve_Word_8 : Word;
      Reserve_Word_10 : Word;
      MC_Place_Number : Byte;
      Mould_Number : Byte;
      Time_Nummer : Byte;
      Offset_of_Shottime : Byte;
      Stepnumber : Byte;   // Schrittmerker für die Ablaufsteuerung der Roboteransteuerung
      Input : "ABB_IRC5_Input";   // Merkerbereich für die Eingänge vom Roboter
      Output : "ABB_IRC5_Output";   // Merkerbereich für die Ausgänge vom Roboter
      Meldungen : "ABB_IRC5_Messages";   // Merkerbereich für die Meldungen vom Roboter
   END_STRUCT;
END_TYPE

TYPE "UDT114_IF_externalPlant"
TITLE = Signals interface external plant
VERSION : 0.1
   STRUCT
      FaultLevel_1 : Bool;   // A fault group 1 exist
      FaultLevel_2 : Bool;   // A fault group 2 exist
      FaultLevel_3 : Bool;   // A fault group 3 exist
      Message_activ : Bool;   // A message is active
      Spare_05 : Bool;
      Spare_06 : Bool;
      Spare_07 : Bool;
      Spare_08 : Bool;
      IF_is_selected : Bool;   // Valid interface data detected and start foaming cycle
      Start_to_Cycle : Bool;   // Pulse to start foaming cycle
      Stop_to_Cycle : Bool;   // Pulse to stop foaming cycle
      HF_StrobeStart : Bool;   // Helping flag of raising edge strobe or start signal
      Spare_13 : Bool;
      FHF_Cycle_Release : Bool;   // Helping flag to set "Strobe" fault
      StatShotOffafterCycleFinish : Bool;   // The start shot signal was "0" after shot finish
      CycleOffafterShotFinish : Bool;   // The cycle was off after shot finish
      PU_ok : Bool;   // Signal to external plant from foaming machine ready for production
      PU_Cycle_runs : Bool;   // Signal to external plant from foaming machine foaming cycle running
      PU_Pouringrelease : Bool;   // Signal to external plant from foaming machine release open mixinghead
      PU_Shotend : Bool;   // Signal to external plant from foaming machine foaming finished
      ExtP_in_Automatic : Bool;   // Signal from external plant at automatic mode
      ExtP_MH_open : Bool;   // Signal from external plant open mixing head
      ExtP_CP_forward : Bool;   // Signal from external plant move cleaning piston mixinghead in front position
      Spare_2_7 : Bool;
      PrgNo_Storage : Byte;   // Program number read in by strobe or start signal
      PrgNo_to_PU : Byte;
      "Step" : Byte;   // Steps of interface program
   END_STRUCT;
END_TYPE

TYPE "UDT115_Test"
TITLE = Signals of discharging by test valves
VERSION : 0.0
   STRUCT
      Test_runs : Bool;   // Ein Zyklus zum Testen der Austragsleistung wurde gestartet
      Test_K1 : Bool;   // Ein Zyklus zum Testen der Austragsleistung der Komponente 1 wurde gestartet
      Test_K2 : Bool;   // Ein Zyklus zum Testen der Austragsleistung der Komponente 2 wurde gestartet
      Test_K3 : Bool;   // Ein Zyklus zum Testen der Austragsleistung der Komponente 3 wurde gestartet
      Test_K4 : Bool;   // Ein Zyklus zum Testen der Austragsleistung der Komponente 4 wurde gestartet
      Start_to_Cycle : Bool;   // Signal zum Starten des Zyklusses zum Testen der Austragsleistung
      Stop_to_Cycle : Bool;   // Signal zum Unterbrechen des Zyklusses zum Testen der Austragsleistung
      Spare_0_7 : Bool;
      Spare_Byte : Byte;
   END_STRUCT;
END_TYPE

TYPE "UDT116_GBE"
TITLE = State of GBE unit
VERSION : 0.1
   STRUCT
      EmergencyStop : Bool;
      FLT_Supply : Bool;
      FLT_Interface : Bool;
      State03 : Bool;
      State04 : Bool;
      State05 : Bool;
      State06 : Bool;
      State07 : Bool;
      GBE_OK : Bool;
      State09 : Bool;
      State10 : Bool;
      State11 : Bool;
      State12 : Bool;
      State13 : Bool;
      State14 : Bool;
      State15 : Bool;
   END_STRUCT;
END_TYPE

TYPE "UDT117_RinsingStation"
TITLE = State of rinsing station, flushing mh and tubes
VERSION : 0.0
   STRUCT
      Warning_Min_Level : Bool;   // Warnung: Der min. Füllstand des Wassertanks wurde unterschritten
      FLT_Min_Level : Bool;   // Störung: Der min. Füllstand des Wassertanks wurde unterschritten (> 5 min.)
      Warning_Min_Temp : Bool;   // Warnung: Die min. Temperatur des Wassertanks wurde unterschritten
      FLT_Min_Temp : Bool;   // Störung: Die min. Temperatur des Wassertanks wurde unterschritten (> 5 min.)
      FLT_Min_Pressure : Bool;   // Störung: Der minimale Reinigungsdruck wurde nicht erreicht
      FLT_Max_Pressure : Bool;   // Störung: Der maximale Reinigungsdruck wurde erreicht
      FLT_SystemAirPressure : Bool;   // Störung: Der minimale Systemluftdruck wurde unterschritten
      FLT_TimeValue_Null : Bool;   // Störung: Die eingegebene Zeitwerte für den Sprühkopf ist = 0
      Step_01 : Bool;   // Open circulation valve component
      Step_02 : Bool;   // Shut valve comonent (2)
      Step_03 : Bool;   // Open valve rinsing agent (3)
      Step_04 : Bool;   // Lock valve rinsing agent open (4)
      Step_05 : Bool;   // Start rinsing pump (5)
      Step_06 : Bool;   // Stop rinsing pump (6)
      Step_07 : Bool;   // Lock valve rinsing agent close (7)
      Step_08 : Bool;   // Start blow air (8)
      CleaningActive : Bool;   // Die Reinigung des Mischkopfes wurde gestartet und läuft
      MH_was_open : Bool;   // Information das der Mischkopf offen war und gereinigt werden muß
      CleanerReady : Bool;   // Der Mischkopfreiniger ist betriebsbereit
      SwitchCleaning_ON_OFF : Bool;   // Signal zum Starten des Mischkopfreinigers
      CleaningFinished : Bool;   // Der Reinigungszyklus des Mischkopfreinigers ist beendet
      BlowAir_OnOFF_manual : Bool;   // Blasluft einschalten von Hand durch Taster
      Rinsing_OnOFF_manual : Bool;   // Spühlmittel einschalten von Hand durch Taster
      FLT_RinsingPump : Bool;   // Fault: Motorprotection rising pump
      Spare_3_0 : Bool;   // --------------
      RinsingPump : Bool;   // Ansteuerung der Spülpumpe zum Reinigen
      Valve_RelRinsingAgent : Bool;   // Ansteuerung der Freigabe für das Spülmittel
      Valve_RinsingAgent : Bool;   // Valve pre run and backflow rinsing agent
      Valve_BlowAir : Bool;   // Ansteuerung der Freigabe für die Blasluft
      ValveComponent : Bool;   // Valve pre run and backflow component
      Spare_3_6 : Bool;   // --------------
      ValveCircComponent : Bool;   // --------------
      StepNumber : Byte;   // Schrittmerker für die Ablaufsteuerung des Mischkopfreinigers
      Interval : Bool;
      doBlowAir : Bool;   // Blasluft ein (von Roboter)
      Pause : Bool;   // --------------
      Step_09 : Bool;   // Shut valve rinsing agent (9)
      Step_10 : Bool;   // Open valve comonent (10)
      Step_11 : Bool;   // Close circulation valve component (11)
      Spare_5_6 : Bool;
      Spare_5_7 : Bool;   // --------------
      StateCleaning : Int;   // 1->BlowAir ON; 2->Fault BlowAir; 3->BlowAir requested but not on
   END_STRUCT;
END_TYPE

TYPE "UDT118_MH_Cleaner"
TITLE = State of mixing head cleaning unit
VERSION : 0.0
   STRUCT
      Warnung_Min_Level : Bool;   // Warnung: Der min. Füllstand des Wassertanks wurde unterschritten
      Stoerung_Min_Level : Bool;   // Störung: Der min. Füllstand des Wassertanks wurde unterschritten (> 5 min.)
      Warnung_Min_Temp : Bool;   // Warnung: Die min. Temperatur des Wassertanks wurde unterschritten
      Stoerung_Min_Temp : Bool;   // Störung: Die min. Temperatur des Wassertanks wurde unterschritten (> 5 min.)
      Stoerung_Heizung : Bool;   // Störung: Der Sicherung oder des Motorschutzes für die Heizung des Wassertanks
      Meldung_Deckel_offen : Bool;   // Meldung: Das der Deckel des Reiniger noch geöffnet ist
      LFI_Zeit_gleich_Null : Bool;   // Störung: Die eingegebene Spül- oder Trocknen- Zeit für den LFI Kopf ist = 0
      SPK_Zeit_gleich_Null : Bool;   // Störung: Die eingegebene Spül- oder Trocknen- Zeit für den Sprühkopf ist = 0
      Stoerung_Max_Level : Bool;   // Störung: Der max. Füllstand des Wassertanks wurde überschritten
      STG_Motorschutz : Bool;   // Störung: Motorschutzschalter
      STG_Trockenlaufschutz : Bool;   // Störung: Trockenlaufschutz der Hochdruckpumpe
      Reserve_1_3 : Bool;
      Reserve_1_4 : Bool;
      Reserve_1_5 : Bool;
      Reserve_1_6 : Bool;
      Reserve_1_7 : Bool;
      MK_Reinigung_Laeuft : Bool;   // Die Reinigung des Mischkopfes wurde gestartet und läuft
      MK_war_offen : Bool;   // Information das der Mischkopf offen war und gereinigt werden muß
      MK_Reiniger_oK : Bool;   // Der Mischkopfreiniger ist betriebsbereit
      MK_Reiniger_start : Bool;   // Signal zum Starten des Mischkopfreinigers
      MK_Reiniger_ende : Bool;   // Der Reinigungszyklus des Mischkopfreinigers ist beendet
      Anforderung_HD_Pumpe : Bool;   // Anforderung der Hochdrucpumpe von extern
      Reserve_2_6 : Bool;   // Fregabe Hochdruckpumpe für extern
      Reserve_2_7 : Bool;
      Kreislaufpumpe : Bool;   // Ansteuerung der Kreislaufpumpe zum Spülen der Wasserführung
      Spuelpumpe : Bool;   // Ansteuerung der Spülpumpe und der gedrosselter Luft zum Reinigen
      Trockenluft : Bool;   // Ansteuerung der Luft zum Trocknen des Mischkopfes
      Ventil_Dichtung : Bool;   // Ansteuerung der Dichtlippe zum Spritzschutz beim Reinigen
      Heizung : Bool;   // Ansteuerung der Heizung zum Aufheizen des Reinigungswassers
      HD_Pumpe_Ein : Bool;   // Ansteuerung Motor Hochdruckpumpe für Sprühkopf
      Ventil_HD_Pumpe : Bool;   // Ansteuerung Ventil Hochdruckpumpe für Sprühkopf
      Reserve_3_7 : Bool;
      Schrittnummer : Byte;   // Schrittmerker für die Ablaufsteuerung des Mischkopfreinigers
      Reserve_5 : Byte;
   END_STRUCT;
END_TYPE

TYPE "UDT119_Bandfilter"
VERSION : 0.0
   STRUCT
      Stoerung_Motorschutz : Bool;   // Störung: Der Sicherung oder des Motorschutzes für den Fließantrieb
      Stoerung_Flies : Bool;   // Störung: Das kein Fließ mehr vorhanden ist
      Stoerung_Zaehler : Bool;   // Störung: Der eingegebene Wert für die Schußzahl ist 0
      Meldung_Deckel_offen : Bool;   // Meldung: Der Deckel des Reiniger ist noch geöffnet
      Reserve_0_4 : Bool;
      Reserve_0_5 : Bool;
      Reserve_0_6 : Bool;
      Reserve_0_7 : Bool;
      Flankenmerker : Bool;   // Flankenmerker zum aufsummieren der Schußanzahl
      Zaehlimpuls : Bool;   // Impulsmerker zum aufsummieren der Schußanzahl
      Vorschub_Automatisch : Bool;   // Der Fließvorschub soll automatisch angesteuert werden (nach Anzahl Schüßen)
      Reserve_1_3 : Bool;
      Reserve_1_4 : Bool;
      Reserve_1_5 : Bool;
      Reserve_1_6 : Bool;
      Vorschub : Bool;   // Ansteuerung des Vorschub- Antriebes
   END_STRUCT;
END_TYPE

TYPE "UDT112_IF_UP_MC"
TITLE = Signals user panel MH, interface mould carrier
VERSION : 0.0
   STRUCT
      FaultLevel_1 : Bool;   // A fault group 1 exist
      FaultLevel_2 : Bool;   // A fault group 2 exist
      FaultLevel_3 : Bool;   // A fault group 3 exist
      Message_activ : Bool;   // A message is active
      IF_is_Selected : Bool;   // The interface is registered for the next foaming cycle
      IF_is_on_1_Position : Bool;   // The interface is at first position at the FIFO
      IF_is_on_2_Position : Bool;   // The interface is at second position at the FIFO
      Start_to_Cycle : Bool;   // Signal to start foaming cycle at this interface
      Stop_to_Cycle : Bool;   // Signal to stop foaming cycle at this interface
      FHF_Fault : Bool;   // Edge flag to built thr interface fault signal
      Shotsend_IF : Bool;   // During interface is at first postion a foaming cycle finished
      Fault_IF : Bool;   // During interface is at first postion a fault occured
      HF_Release_IF : Bool;   // Edge flag to build the signal to register the interface
      Stop_Buton_switched : Bool;   // Helpflag of a recognition of the stop button at FIFO- Position > 2
      FHF_KLZ2 : Bool;   // Edge flag to build the shot end signal during KLZ2
      HF_T_Start_MH : Bool;   // Edge flag to build the signal whne "Start MH" button is pressed
   END_STRUCT;
END_TYPE

TYPE "UDT121_DF_Chanel"
TITLE = State and index of a flow channel
VERSION : 0.0
   STRUCT
      OUT_PROCAN : Struct   // Signals from plc to proc module
         FlowIndex : Struct
            FlowIndex0 : Bool;
            FlowIndex1 : Bool;
            FlowIndex2 : Bool;
            FlowIndex3 : Bool;
            Spare4 : Bool;
            Notclosedloop : Bool;   // flow is not closed loop controlled
            StartQPB : Bool;   // toggle flag: start FPB now
            Enableclosedloop : Bool;   // Enable close loop control
         END_STRUCT;
         TandemComand : Word;
         SpareWord : Word;
         Spare_DWORD_56 : DWord;
      END_STRUCT;
      IN_PROCAN : Struct   // Signals from proc module to plc
         Flowrate : DInt;
         PistonPosition : DInt;
         TandemStatus : Word;
         Flow_Status : Struct
            Flowstopped : Bool;   // piston has stopped
            FlowQPB : Bool;   // Flow quick pressure build up is active
            ControlOnUpperLimit : Bool;   // flow control loop operates on it upper limits
            ControlOnLowerLimit : Bool;   // flow control loop operates on its lower limits
            FlowtoleranceL : Bool;   // tolerance: flow is too low
            FlowtoleranceH : Bool;   // tolerance: flow is too high
         END_STRUCT;
         Spare_DWORD_96 : DWord;
      END_STRUCT;
   END_STRUCT;
END_TYPE

TYPE "UDT100_EdgeFilter"
TITLE = State of auxiliary drive
VERSION : 0.0
   STRUCT
      FLT_Exist : Bool;
      FaultLevel_3 : Bool;   // A fault group 3 exist
      Reset_Intervall : Bool;   // Reset of intervall- mode at running- and pausetime
      Run : Bool;   // Drive at intervall- mode in running
      Pause : Bool;   // Drive at intervall- mode in pause time
      Spare_6 : Bool;
      Spare_7 : Bool;
      Spare_8 : Bool;
      Spare_9 : Bool;
      Spare_10 : Bool;
      Spare_11 : Bool;
      Spare_12 : Bool;
      Spare_13 : Bool;
      Spare_14 : Bool;
      Spare_15 : Bool;
      Switch_Drive_ON_OFF : Bool;   // Switch auxiliary drive ON-OFF (external signal)
      State_Drive : Int;   // 1->Drive ON; 2->Fault Drive; 3->Drive requested but not on
   END_STRUCT;
END_TYPE

TYPE "UDT123_MH_Chanel"
TITLE = State and control signals of steering piston
VERSION : 0.0
   STRUCT
      IN : Struct
         MH_With_CleaningPiston : Bool;
         MH_EmergencyStop : Bool;
         MH_APS_CleaningPiston : Bool;   // Approximate switch cleaning piston
         MH_Aps_Mixinghead : Bool;   // Approximate switch steering piston
         MH_Release_SWU : Bool;
         MH_Manual_Mode : Bool;
         MH_Auto_Mode : Bool;
         MH_Prep_Foaming_MC : Bool;
         MH_Releas_Foaming_MC : Bool;
         MH_HP_Circ_MH : Bool;
         MH_Start : Bool;
         MH_Stop : Bool;
         MH_CP_forward : Bool;
         MH_CP_backward : Bool;
         Spare_1_6 : Bool;
         Spare_1_7 : Bool;
         MH_Prog_No_MH : Byte;
         Shottime : Real;
         MH_Opentime : Real;
         MH_Closingtime : Real;
         MH_Status : Struct
            NoShotReleaseFromCP : Bool;
            NoShotReleaseFromExtern : Bool;
            Ready4Shot : Bool;
            shotactive_MH : Bool;
            shotdone_MH : Bool;
            Spare5 : Bool;
            Spare6 : Bool;
            Spare7 : Bool;
            SPFopening_MH : Bool;
            SPFclosing_MH : Bool;
            SPFopen_MH : Bool;
            SPFclosed_MH : Bool;
            MHBouncing : Bool;
            SPFaborted_SoftwareRelease : Bool;
            SPFaborted_CP : Bool;
            SPFabortet_HardwareRelease : Bool;
         END_STRUCT;
         PLC_State : Int;
         CleaningPistonState : Struct
            CP_to_slow_FW_MH : Bool;   // CP moves too slow forward
            CP_to_slow_BW_MH : Bool;   // CP moves too slow back
            CP_MovesDuringShot_MH : Bool;   // CP moves during shot
            CP_DontReachFWPos_MH : Bool;
            CP_DontReachBWPos_MH : Bool;
            CP_LeaveHP_MH : Bool;
            CP_inFWPosition_MH : Bool;   // CP is in front position
            CP_inBWPosition_MH : Bool;   // CP is back (ready for shot)
         END_STRUCT;
      END_STRUCT;
      OUT : Struct
         MH : Struct
            V_SWU_MH : Bool;   // Valve switch over unit
            H_Shotcounter_MH : Bool;   // indicator shot counter
            V_CP_Forward_MH : Bool;   // Valve cleaning piston forward
            H_CP_Back_MH : Bool;   // indicator cleaning piston back
            H_Rel_Foaming_MH : Bool;   // indicator release foaming
            H_HighPressure_MH : Bool;   // indicator high pressure circulation
            K_Fault_MC : Bool;   // malfunction PU-machine to mouldcarrier
            K_ShotEnd_MC : Bool;   // Shotend PU-machine to mouldcarrier
            V_MH : Bool;   // Valve mixinghead open
            spare11 : Bool;
            spare12 : Bool;
            spare13 : Bool;
            spare14 : Bool;
            spare15 : Bool;
            spare16 : Bool;
            V_LowPressure_Circ_MH : Bool;   // low pressure circulation
            Shottime : Real;
            ServiceProduction : Int;
         END_STRUCT;
         MH_Control : Struct
            MH_start_shot : Bool;   // shot validation (starts shot with rising edge)
            MH_CP_after_shot : Bool;   // clean after shot (not implemented)
            MH_CP_forward_manual : Bool;   // move CP forward
            MH_Reserve_4 : Bool;
            MH_Reserve_5 : Bool;
            MH_Reserve_6 : Bool;
            MH_Reserve_7 : Bool;
            MH_Reserve_8 : Bool;   // hold shot results
         END_STRUCT;
         PLC_Comand_SP : Byte;
         PLC_Comand_CP : Byte;
         PLC_Set_Value_SP : Int;
         PLC_Set_Value_CP : Int;
         NozzelBypassControl : Word;
         NozzelBypassSetOut : Word;
      END_STRUCT;
      MH_Ref_OK : Bool;
      MH_INI : Bool;
      CP_INI : Bool;
      V_Nozzel01 : Bool;
      V_Nozzel02 : Bool;
      V_MH : Bool;
      Spare06 : Bool;
      Spare07 : Bool;
   END_STRUCT;
END_TYPE

